
       #AUX_rgtSendBuffer.dLung := 0;
       #AUX_rgtSendBuffer.dID := #AUX_rgtSendBuffer.dID + 1;
       #AUX_rgtSendBuffer.dThick_um := #INO_tTrack.tLastPlacedCap.dThick_cmm;
   //    WRITE_BIG(src_variable := _byte_in_, dest_array := _variant_inout_, pos := _dint_inout_);
       #TMP_dPos := 0;
       #TMP_iRetVal:= WRITE_LITTLE(src_variable :=  #AUX_rgtSendBuffer.dLung, dest_array :=  #AUX_rgtSendBuffer_LittleEndian, pos := #TMP_dPos);
       #TMP_dPos := 4;
       #TMP_iRetVal := WRITE_LITTLE(src_variable := #AUX_rgtSendBuffer.dID, dest_array := #AUX_rgtSendBuffer_LittleEndian, pos := #TMP_dPos);
       #TMP_dPos := 8;
       #TMP_iRetVal := WRITE_LITTLE(src_variable := #AUX_rgtSendBuffer.dThick_um, dest_array := #AUX_rgtSendBuffer_LittleEndian, pos := #TMP_dPos);
       #AUX_dNumByteToSend := 0;
   END_IF;
END_REGION

REGION Network 25: ### SEND DATA TO CAMERA
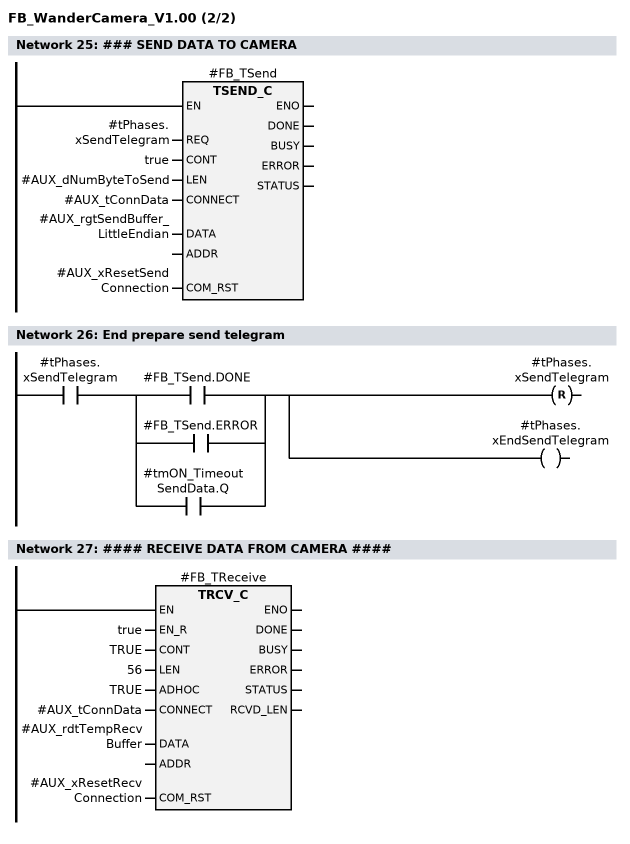
   #FB_TSend(REQ := #tPhases.xSendTelegram,   // TSEND_C
             CONT := true,
             LEN := #AUX_dNumByteToSend,
             CONNECT := #AUX_tConnData,
             DATA := #AUX_rgtSendBuffer_LittleEndian,
             COM_RST := #AUX_xResetSendConnection);
END_REGION

REGION Network 26: End prepare send telegram
   RUNG wire#powerrail
      Contact( #tPhases.xSendTelegram )
      wire#w1
      Contact( #FB_TSend.DONE )
      wire#w2
      R_Coil( #tPhases.xSendTelegram )
   END_RUNG
   RUNG wire#w1
      Contact( #FB_TSend.ERROR )
   END_RUNG wire#w2
   RUNG wire#w1
      Contact( #tmON_TimeoutSendData.Q )
   END_RUNG wire#w2
   RUNG wire#w2
      Coil( #tPhases.xEndSendTelegram )
   END_RUNG
   // the same network as SCL:
   #_w1 := #tPhases.xSendTelegram AND (#FB_TSend.DONE OR #FB_TSend.ERROR OR #tmON_TimeoutSendData.Q);
   IF #_w1 THEN #tPhases.xSendTelegram := FALSE; END_IF;
   #tPhases.xEndSendTelegram := #_w1;
END_REGION

REGION Network 27: #### RECEIVE DATA FROM CAMERA ####
   #FB_TReceive(EN_R := true,   // TRCV_C
                CONT := TRUE,
                LEN := 56,
                ADHOC := TRUE,
                CONNECT := #AUX_tConnData,
                DATA := #AUX_rdtTempRecvBuffer,
                COM_RST := #AUX_xResetRecvConnection);
END_REGION

REGION Network 28 (SCL): Manage data received
   IF #FB_TReceive.DONE THEN

       IF #FB_TReceive.RCVD_LEN > 0 THEN
           #TMP_dPos := 0;
           #TMP_iRetVal:= READ_LITTLE(src_array:=#AUX_rdtTempRecvBuffer, dest_Variable=>#AUX_rdtRecvBuffer.dLung, pos:=#TMP_dPos);
           #TMP_dPos := 4;
           #TMP_iRetVal := READ_LITTLE(src_array := #AUX_rdtTempRecvBuffer, dest_Variable => #AUX_rdtRecvBuffer.dID, pos := #TMP_dPos);
           #TMP_dPos := 8;
           #TMP_iRetVal := READ_LITTLE(src_array := #AUX_rdtTempRecvBuffer, dest_Variable => #AUX_rdtRecvBuffer.dTime1, pos := #TMP_dPos);
           #TMP_dPos := 12;
           #TMP_iRetVal := READ_LITTLE(src_array := #AUX_rdtTempRecvBuffer, dest_Variable => #AUX_rdtRecvBuffer.dTime2, pos := #TMP_dPos);
           #TMP_dPos := 16;
           #TMP_iRetVal := READ_LITTLE(src_array := #AUX_rdtTempRecvBuffer, dest_Variable => #AUX_rdtRecvBuffer.dStato, pos := #TMP_dPos);
           #TMP_dPos := 20;
           #TMP_iRetVal := READ_LITTLE(src_array := #AUX_rdtTempRecvBuffer, dest_Variable => #AUX_rdtRecvBuffer.dGrossZeroSide_um, pos := #TMP_dPos);
           #TMP_dPos := 24;
           #TMP_iRetVal := READ_LITTLE(src_array := #AUX_rdtTempRecvBuffer, dest_Variable => #AUX_rdtRecvBuffer.dNetExtZeroSide_um, pos := #TMP_dPos);
           #TMP_dPos := 28;
           #TMP_iRetVal := READ_LITTLE(src_array := #AUX_rdtTempRecvBuffer, dest_Variable => #AUX_rdtRecvBuffer.dNetCenterZeroSide_um, pos := #TMP_dPos);
           #TMP_dPos := 32;
           #TMP_iRetVal := READ_LITTLE(src_array := #AUX_rdtTempRecvBuffer, dest_Variable => #AUX_rdtRecvBuffer.dNetZeroSide_um, pos := #TMP_dPos);
           #TMP_dPos := 36;
           #TMP_iRetVal := READ_LITTLE(src_array := #AUX_rdtTempRecvBuffer, dest_Variable => #AUX_rdtRecvBuffer.dGrossOppSide_um, pos := #TMP_dPos);
           #TMP_dPos := 40;
           #TMP_iRetVal := READ_LITTLE(src_array := #AUX_rdtTempRecvBuffer, dest_Variable => #AUX_rdtRecvBuffer.dNetExtOppoSide_um, pos := #TMP_dPos);
           #TMP_dPos := 44;
           #TMP_iRetVal := READ_LITTLE(src_array := #AUX_rdtTempRecvBuffer, dest_Variable => #AUX_rdtRecvBuffer.dNetCenterOppoSide_um, pos := #TMP_dPos);
           #TMP_dPos := 48;
           #TMP_iRetVal := READ_LITTLE(src_array := #AUX_rdtTempRecvBuffer, dest_Variable => #AUX_rdtRecvBuffer.dNetOppoSide_um, pos := #TMP_dPos);
           #TMP_dPos := 52;
           #TMP_iRetVal := READ_LITTLE(src_array := #AUX_rdtTempRecvBuffer, dest_Variable => #AUX_rdtRecvBuffer.dLength, pos := #TMP_dPos);

           #OS_xNewDataAvailable := 1;
           #INO_tRibbon.rgtGlassData[#IN_dGlassDataMachineIndex].dDistSnapRoll_cmm := #tHMR.dDistanceFromSnaproll_cmm;

           //Update the position
           IF NOT #INO_tRibbon.rgtGlassDataUpdate[#IN_dGlassDataMachineIndex].xUpdateRequest THEN
               #INO_tRibbon.rgtGlassDataUpdate[#IN_dGlassDataMachineIndex].tData.dGrossWander_cmm := #tHMR.dCurrentGrossWander_cmm;
               #INO_tRibbon.rgtGlassDataUpdate[#IN_dGlassDataMachineIndex].tData.dNetWander_cmm := #tHMR.dCurrentNetWander_cmm;
               #INO_tRibbon.rgtGlassDataUpdate[#IN_dGlassDataMachineIndex].tData.dGrossWidth_cmm := #tHMR.dCurrentGrossWidth_cmm;
               #INO_tRibbon.rgtGlassDataUpdate[#IN_dGlassDataMachineIndex].tData.dNetWidth_cmm := #tHMR.dCurrentNetWidth_cmm;
               #INO_tRibbon.rgtGlassDataUpdate[#IN_dGlassDataMachineIndex].xUpdateRequest := TRUE;
           END_IF;
       END_IF;

   END_IF;
END_REGION

REGION Network 29 (SCL): Phase in progress
   GATHER(IN:=#tPhases,
          OUT=>#TMP_dwValue);

   IF #TMP_dwValue <> 0 THEN
       #ST_xPhaseProgr := TRUE;
   ELSE
       #ST_xPhaseProgr := FALSE;
   END_IF;
END_REGION
END_FUNCTION_BLOCK

// folder: 03_Programs_Logics/MCC1201/09_Zone

FUNCTION "ZUPS_Faults" : Void   // FC15, LAD
{ S7_Optimized_Access := 'TRUE' }
VERSION : 0.1
   VAR_TEMP
      TMP_dwValue : DWord;
   END_VAR
BEGIN

REGION Network 1 (SCL): Reset alarms
   IF "ZUPS".tmOFF_ResetAlarm.OUT_xDone THEN

       #TMP_dwValue := 0;

       SCATTER(IN := #TMP_dwValue,
               OUT => "DB_ZUPS_HMI".tAlm.tE);

       SCATTER(IN := #TMP_dwValue,
               OUT => "DB_ZUPS_HMI".tAlm.tS);

       SCATTER(IN := #TMP_dwValue,
               OUT => "DB_ZUPS_HMI".tAlm.tF);

       SCATTER(IN := #TMP_dwValue,
               OUT => "DB_ZUPS_HMI".tAlm.tW);

   END_IF;
END_REGION

REGION Network 2: Anomalies
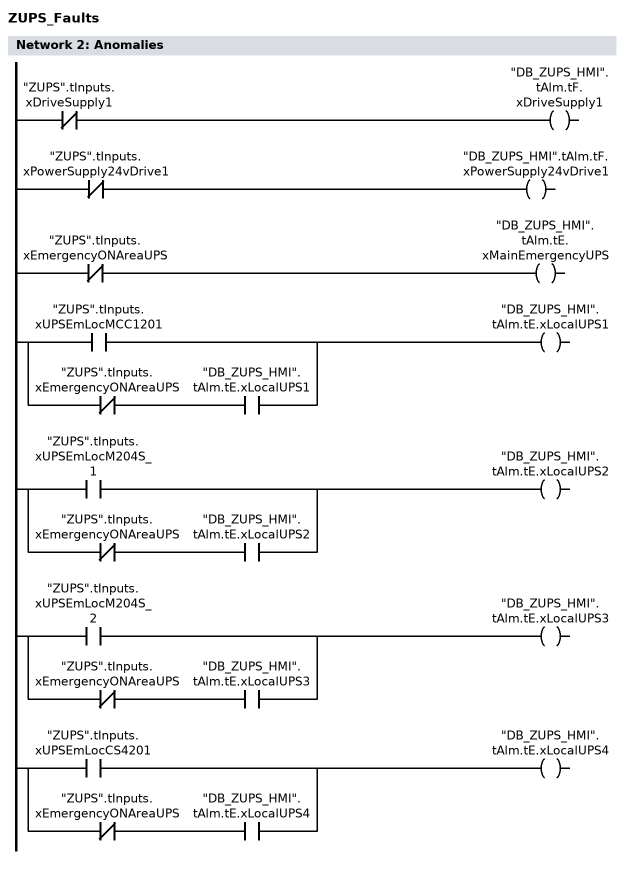
   RUNG wire#powerrail
      I_Contact( "ZUPS".tInputs.xDriveSupply1 )
      Coil( "DB_ZUPS_HMI".tAlm.tF.xDriveSupply1 )
   END_RUNG
   RUNG wire#powerrail
      I_Contact( "ZUPS".tInputs.xPowerSupply24vDrive1 )
      Coil( "DB_ZUPS_HMI".tAlm.tF.xPowerSupply24vDrive1 )
   END_RUNG
   RUNG wire#powerrail
      I_Contact( "ZUPS".tInputs.xEmergencyONAreaUPS )
      Coil( "DB_ZUPS_HMI".tAlm.tE.xMainEmergencyUPS )
   END_RUNG
   RUNG wire#powerrail
      Contact( "ZUPS".tInputs.xUPSEmLocMCC1201 )
      wire#w1
      Coil( "DB_ZUPS_HMI".tAlm.tE.xLocalUPS1 )
   END_RUNG
   RUNG wire#powerrail
      I_Contact( "ZUPS".tInputs.xEmergencyONAreaUPS )
      Contact( "DB_ZUPS_HMI".tAlm.tE.xLocalUPS1 )
   END_RUNG wire#w1
   RUNG wire#powerrail
      Contact( "ZUPS".tInputs.xUPSEmLocM204S_1 )
      wire#w2
      Coil( "DB_ZUPS_HMI".tAlm.tE.xLocalUPS2 )
   END_RUNG
   RUNG wire#powerrail
      I_Contact( "ZUPS".tInputs.xEmergencyONAreaUPS )
      Contact( "DB_ZUPS_HMI".tAlm.tE.xLocalUPS2 )
   END_RUNG wire#w2
   RUNG wire#powerrail
      Contact( "ZUPS".tInputs.xUPSEmLocM204S_2 )
      wire#w3
      Coil( "DB_ZUPS_HMI".tAlm.tE.xLocalUPS3 )
   END_RUNG
   RUNG wire#powerrail
      I_Contact( "ZUPS".tInputs.xEmergencyONAreaUPS )
      Contact( "DB_ZUPS_HMI".tAlm.tE.xLocalUPS3 )
   END_RUNG wire#w3
   RUNG wire#powerrail
      Contact( "ZUPS".tInputs.xUPSEmLocCS4201 )
      wire#w4
      Coil( "DB_ZUPS_HMI".tAlm.tE.xLocalUPS4 )
   END_RUNG
   RUNG wire#powerrail
      I_Contact( "ZUPS".tInputs.xEmergencyONAreaUPS )
      Contact( "DB_ZUPS_HMI".tAlm.tE.xLocalUPS4 )
   END_RUNG wire#w4
   // the same network as SCL:
   "DB_ZUPS_HMI".tAlm.tF.xDriveSupply1 := NOT "ZUPS".tInputs.xDriveSupply1;
   "DB_ZUPS_HMI".tAlm.tF.xPowerSupply24vDrive1 := NOT "ZUPS".tInputs.xPowerSupply24vDrive1;
   "DB_ZUPS_HMI".tAlm.tE.xMainEmergencyUPS := NOT "ZUPS".tInputs.xEmergencyONAreaUPS;
   "DB_ZUPS_HMI".tAlm.tE.xLocalUPS1 := "ZUPS".tInputs.xUPSEmLocMCC1201 OR (NOT "ZUPS".tInputs.xEmergencyONAreaUPS AND "DB_ZUPS_HMI".tAlm.tE.xLocalUPS1);
   "DB_ZUPS_HMI".tAlm.tE.xLocalUPS2 := "ZUPS".tInputs.xUPSEmLocM204S_1 OR (NOT "ZUPS".tInputs.xEmergencyONAreaUPS AND "DB_ZUPS_HMI".tAlm.tE.xLocalUPS2);
   "DB_ZUPS_HMI".tAlm.tE.xLocalUPS3 := "ZUPS".tInputs.xUPSEmLocM204S_2 OR (NOT "ZUPS".tInputs.xEmergencyONAreaUPS AND "DB_ZUPS_HMI".tAlm.tE.xLocalUPS3);
   "DB_ZUPS_HMI".tAlm.tE.xLocalUPS4 := "ZUPS".tInputs.xUPSEmLocCS4201 OR (NOT "ZUPS".tInputs.xEmergencyONAreaUPS AND "DB_ZUPS_HMI".tAlm.tE.xLocalUPS4);
END_REGION

REGION Network 3 (SCL): Calculate comulative status
   GATHER(IN:="DB_ZUPS_HMI".tAlm.tE,
              OUT=>#TMP_dwValue);

       IF "DB_ZUPS_HMI".tAlm.tE.xMainEmergencyUPS THEN
       "ZUPS".ST_xZoneEmergency := TRUE;
   ELSE
       "ZUPS".ST_xZoneEmergency := FALSE;
   END_IF;

   GATHER(IN:="DB_ZUPS_HMI".tAlm.tS,
              OUT=>#TMP_dwValue);

   IF #TMP_dwValue <> 0 THEN
       "ZUPS".ST_xZoneStoppingFaults := TRUE;
   ELSE
       "ZUPS".ST_xZoneStoppingFaults := FALSE;
   END_IF;

   GATHER(IN:="DB_ZUPS_HMI".tAlm.tF,
              OUT=>#TMP_dwValue);

   IF #TMP_dwValue <> 0 THEN
       "ZUPS".ST_xZoneFaults := TRUE;
   ELSE
       "ZUPS".ST_xZoneFaults := FALSE;
   END_IF;

   GATHER(IN:="DB_ZUPS_HMI".tAlm.tW,
              OUT=>#TMP_dwValue);

   IF #TMP_dwValue <> 0 THEN
       "ZUPS".ST_xZoneWarnings := TRUE;
   ELSE
       "ZUPS".ST_xZoneWarnings := FALSE;
   END_IF;

   IF "ZUPS".ST_xZoneEmergency AND "ZUPS".ST_xZoneStoppingFaults AND "ZUPS".ST_xZoneFaults THEN
       "ZUPS".ST_xZoneError := TRUE;
   ELSE
       "ZUPS".ST_xZoneError := FALSE;
   END_IF;
END_REGION
END_FUNCTION

FUNCTION "ZUPS_Logics" : Void   // FC17, LAD
{ S7_Optimized_Access := 'TRUE' }
VERSION : 0.1
   VAR_TEMP
      TMP_rlVal : LReal;
   END_VAR
   VAR_TEMP   // added for the SCL form of the ladder/FBD networks
      _w1 : Bool;
      _w2 : Bool;
   END_VAR
BEGIN

REGION Network 1: #### CONSTANTS ####
END_REGION

REGION Network 2 (SCL): ### SIMULATION ###
   IF "SIMULATION_ACTIVE" THEN
       "ZUPS".tInputs.xDriveSupply1 := TRUE;
       "ZUPS".tInputs.xPowerSupply24vDrive1 := TRUE; 
       "ZUPS".tInputs.xEmergencyONAreaUPS := true;

   END_IF;
END_REGION

REGION Network 3: #### MATCH ####
END_REGION

REGION Network 4: Emergency UPS OK delayed
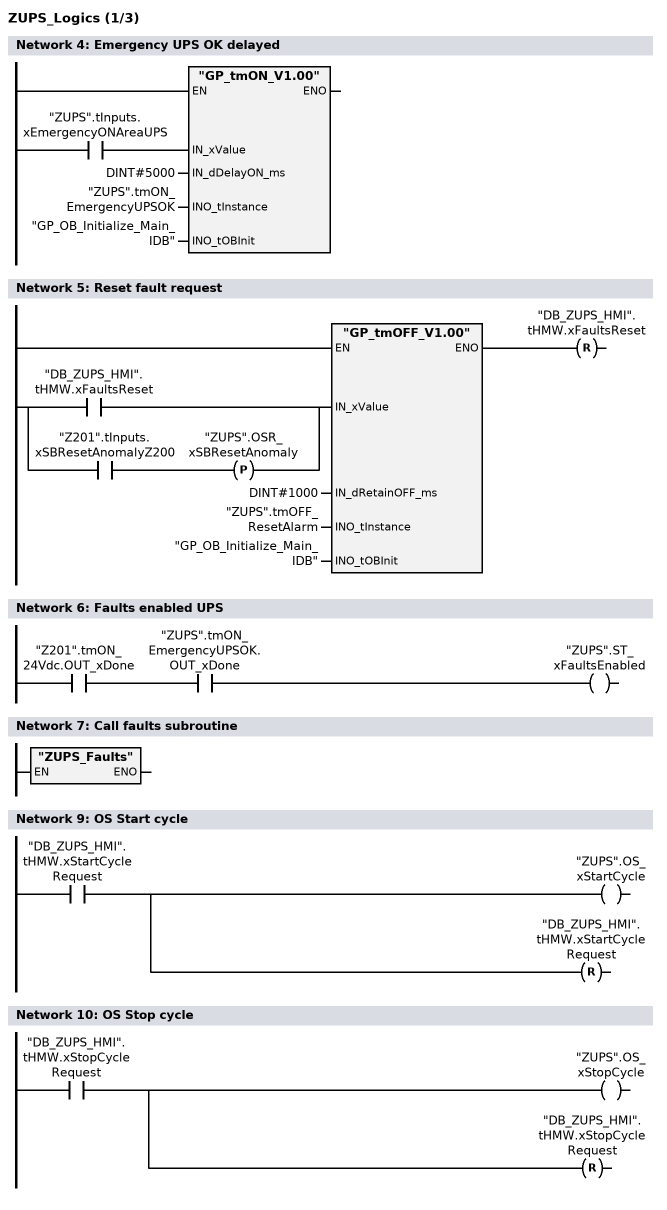
   RUNG wire#powerrail
      "GP_tmON_V1.00"(IN_xValue := wire#w1, IN_dDelayON_ms := DINT#5000, INO_tInstance := "ZUPS".tmON_EmergencyUPSOK, INO_tOBInit := "GP_OB_Initialize_Main_IDB")
   END_RUNG
   RUNG wire#powerrail
      Contact( "ZUPS".tInputs.xEmergencyONAreaUPS )
   END_RUNG wire#w1
   // the same network as SCL:
   "GP_tmON_V1.00"(IN_xValue := "ZUPS".tInputs.xEmergencyONAreaUPS,
                   IN_dDelayON_ms := DINT#5000,
                   INO_tInstance := "ZUPS".tmON_EmergencyUPSOK,
                   INO_tOBInit := "GP_OB_Initialize_Main_IDB");
END_REGION

REGION Network 5: Reset fault request
   RUNG wire#powerrail
      "GP_tmOFF_V1.00"(IN_xValue := wire#w1, IN_dRetainOFF_ms := DINT#1000, INO_tInstance := "ZUPS".tmOFF_ResetAlarm, INO_tOBInit := "GP_OB_Initialize_Main_IDB")
      R_Coil( "DB_ZUPS_HMI".tHMW.xFaultsReset )
   END_RUNG
   RUNG wire#powerrail
      Contact( "DB_ZUPS_HMI".tHMW.xFaultsReset )
   END_RUNG wire#w1
   RUNG wire#powerrail
      Contact( "Z201".tInputs.xSBResetAnomalyZ200 )
      P_Trig( "ZUPS".OSR_xSBResetAnomaly )
   END_RUNG wire#w1
   // the same network as SCL:
   #_w1 := "Z201".tInputs.xSBResetAnomalyZ200 AND NOT "ZUPS".OSR_xSBResetAnomaly;   // rising edge
   "ZUPS".OSR_xSBResetAnomaly := "Z201".tInputs.xSBResetAnomalyZ200;
   "GP_tmOFF_V1.00"(IN_xValue := "DB_ZUPS_HMI".tHMW.xFaultsReset OR #_w1,
                    IN_dRetainOFF_ms := DINT#1000,
                    INO_tInstance := "ZUPS".tmOFF_ResetAlarm,
                    INO_tOBInit := "GP_OB_Initialize_Main_IDB",
                    ENO => #_w2);
   IF #_w2 THEN "DB_ZUPS_HMI".tHMW.xFaultsReset := FALSE; END_IF;
END_REGION

REGION Network 6: Faults enabled UPS
   RUNG wire#powerrail
      Contact( "Z201".tmON_24Vdc.OUT_xDone )
      Contact( "ZUPS".tmON_EmergencyUPSOK.OUT_xDone )
      Coil( "ZUPS".ST_xFaultsEnabled )
   END_RUNG
   // the same network as SCL:
   "ZUPS".ST_xFaultsEnabled := "Z201".tmON_24Vdc.OUT_xDone AND "ZUPS".tmON_EmergencyUPSOK.OUT_xDone;
END_REGION

REGION Network 7: Call faults subroutine
   RUNG wire#powerrail
      "ZUPS_Faults"()
   END_RUNG
   // the same network as SCL:
   "ZUPS_Faults"();
END_REGION

REGION Network 8: #### START/STOP ZONE ####
END_REGION

REGION Network 9: OS Start cycle
   RUNG wire#powerrail
      Contact( "DB_ZUPS_HMI".tHMW.xStartCycleRequest )
      wire#w1
      Coil( "ZUPS".OS_xStartCycle )
   END_RUNG
   RUNG wire#w1
      R_Coil( "DB_ZUPS_HMI".tHMW.xStartCycleRequest )
   END_RUNG
   // the same network as SCL:
   "ZUPS".OS_xStartCycle := "DB_ZUPS_HMI".tHMW.xStartCycleRequest;
   IF "DB_ZUPS_HMI".tHMW.xStartCycleRequest THEN "DB_ZUPS_HMI".tHMW.xStartCycleRequest := FALSE; END_IF;
END_REGION

REGION Network 10: OS Stop cycle
   RUNG wire#powerrail
      Contact( "DB_ZUPS_HMI".tHMW.xStopCycleRequest )
      wire#w1
      Coil( "ZUPS".OS_xStopCycle )
   END_RUNG
   RUNG wire#w1
      R_Coil( "DB_ZUPS_HMI".tHMW.xStopCycleRequest )
   END_RUNG
   // the same network as SCL:
   "ZUPS".OS_xStopCycle := "DB_ZUPS_HMI".tHMW.xStopCycleRequest;
   IF "DB_ZUPS_HMI".tHMW.xStopCycleRequest THEN "DB_ZUPS_HMI".tHMW.xStopCycleRequest := FALSE; END_IF;
END_REGION

REGION Network 11: OS Force stop cycle
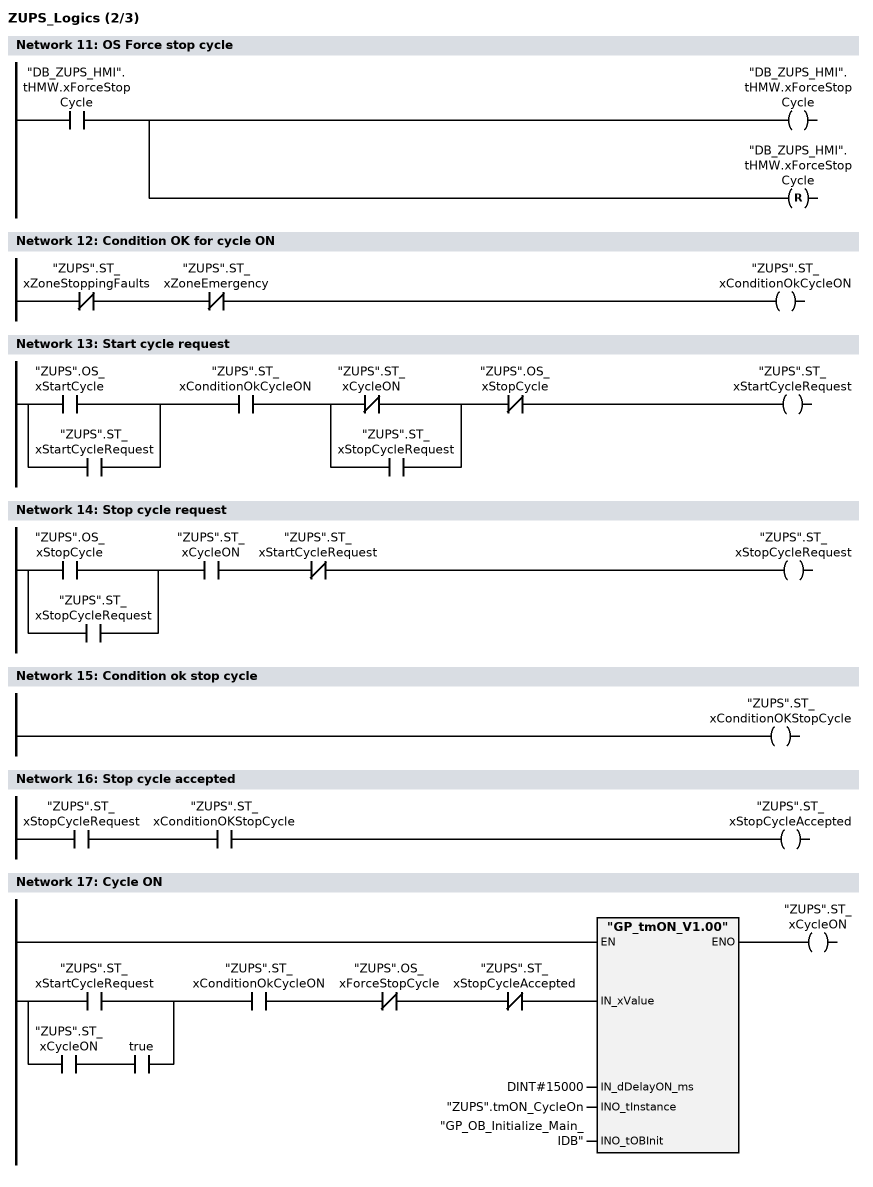
   RUNG wire#powerrail
      Contact( "DB_ZUPS_HMI".tHMW.xForceStopCycle )
      wire#w1
      Coil( "DB_ZUPS_HMI".tHMW.xForceStopCycle )
   END_RUNG
   RUNG wire#w1
      R_Coil( "DB_ZUPS_HMI".tHMW.xForceStopCycle )
   END_RUNG
   // the same network as SCL:
   #_w1 := "DB_ZUPS_HMI".tHMW.xForceStopCycle;
   "DB_ZUPS_HMI".tHMW.xForceStopCycle := "DB_ZUPS_HMI".tHMW.xForceStopCycle;
   IF #_w1 THEN "DB_ZUPS_HMI".tHMW.xForceStopCycle := FALSE; END_IF;
END_REGION

REGION Network 12: Condition OK for cycle ON
   RUNG wire#powerrail
      I_Contact( "ZUPS".ST_xZoneStoppingFaults )
      I_Contact( "ZUPS".ST_xZoneEmergency )
      Coil( "ZUPS".ST_xConditionOkCycleON )
   END_RUNG
   // the same network as SCL:
   "ZUPS".ST_xConditionOkCycleON := NOT "ZUPS".ST_xZoneStoppingFaults AND NOT "ZUPS".ST_xZoneEmergency;
END_REGION

REGION Network 13: Start cycle request
   RUNG wire#powerrail
      Contact( "ZUPS".OS_xStartCycle )
      wire#w1
      Contact( "ZUPS".ST_xConditionOkCycleON )
      wire#w2
      I_Contact( "ZUPS".ST_xCycleON )
      wire#w3
      I_Contact( "ZUPS".OS_xStopCycle )
      Coil( "ZUPS".ST_xStartCycleRequest )
   END_RUNG
   RUNG wire#powerrail
      Contact( "ZUPS".ST_xStartCycleRequest )
   END_RUNG wire#w1
   RUNG wire#w2
      Contact( "ZUPS".ST_xStopCycleRequest )
   END_RUNG wire#w3
   // the same network as SCL:
   "ZUPS".ST_xStartCycleRequest := ("ZUPS".OS_xStartCycle OR "ZUPS".ST_xStartCycleRequest) AND "ZUPS".ST_xConditionOkCycleON AND (NOT "ZUPS".ST_xCycleON OR "ZUPS".ST_xStopCycleRequest) AND NOT "ZUPS".OS_xStopCycle;
END_REGION

REGION Network 14: Stop cycle request
   RUNG wire#powerrail
      Contact( "ZUPS".OS_xStopCycle )
      wire#w1
      Contact( "ZUPS".ST_xCycleON )
      I_Contact( "ZUPS".ST_xStartCycleRequest )
      Coil( "ZUPS".ST_xStopCycleRequest )
   END_RUNG
   RUNG wire#powerrail
      Contact( "ZUPS".ST_xStopCycleRequest )
   END_RUNG wire#w1
   // the same network as SCL:
   "ZUPS".ST_xStopCycleRequest := ("ZUPS".OS_xStopCycle OR "ZUPS".ST_xStopCycleRequest) AND "ZUPS".ST_xCycleON AND NOT "ZUPS".ST_xStartCycleRequest;
END_REGION

REGION Network 15: Condition ok stop cycle
   RUNG wire#powerrail
      Coil( "ZUPS".ST_xConditionOKStopCycle )
   END_RUNG
   // the same network as SCL:
   "ZUPS".ST_xConditionOKStopCycle := TRUE;
END_REGION

REGION Network 16: Stop cycle accepted
   RUNG wire#powerrail
      Contact( "ZUPS".ST_xStopCycleRequest )
      Contact( "ZUPS".ST_xConditionOKStopCycle )
      Coil( "ZUPS".ST_xStopCycleAccepted )
   END_RUNG
   // the same network as SCL:
   "ZUPS".ST_xStopCycleAccepted := "ZUPS".ST_xStopCycleRequest AND "ZUPS".ST_xConditionOKStopCycle;
END_REGION

REGION Network 17: Cycle ON
   RUNG wire#powerrail
      "GP_tmON_V1.00"(IN_xValue := wire#w2, IN_dDelayON_ms := DINT#15000, INO_tInstance := "ZUPS".tmON_CycleOn, INO_tOBInit := "GP_OB_Initialize_Main_IDB")
      Coil( "ZUPS".ST_xCycleON )
   END_RUNG
   RUNG wire#powerrail
      Contact( "ZUPS".ST_xStartCycleRequest )
      wire#w1
      Contact( "ZUPS".ST_xConditionOkCycleON )
      I_Contact( "ZUPS".OS_xForceStopCycle )
      I_Contact( "ZUPS".ST_xStopCycleAccepted )
   END_RUNG wire#w2
   RUNG wire#powerrail
      Contact( "ZUPS".ST_xCycleON )
      Contact( true )
   END_RUNG wire#w1
   // the same network as SCL:
   "GP_tmON_V1.00"(IN_xValue := ("ZUPS".ST_xStartCycleRequest OR ("ZUPS".ST_xCycleON AND true)) AND "ZUPS".ST_xConditionOkCycleON AND NOT "ZUPS".OS_xForceStopCycle AND NOT "ZUPS".ST_xStopCycleAccepted,
                   IN_dDelayON_ms := DINT#15000,
                   INO_tInstance := "ZUPS".tmON_CycleOn,
                   INO_tOBInit := "GP_OB_Initialize_Main_IDB",
                   ENO => #_w1);
   "ZUPS".ST_xCycleON := #_w1;
END_REGION

REGION Network 18: Cycle ON delayed
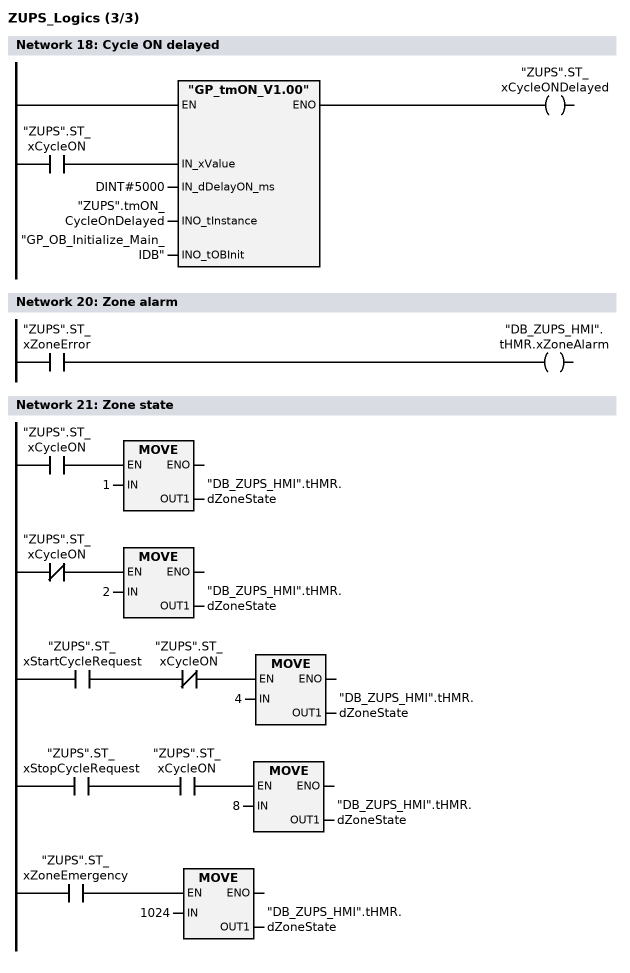
   RUNG wire#powerrail
      "GP_tmON_V1.00"(IN_xValue := wire#w1, IN_dDelayON_ms := DINT#5000, INO_tInstance := "ZUPS".tmON_CycleOnDelayed, INO_tOBInit := "GP_OB_Initialize_Main_IDB")
      Coil( "ZUPS".ST_xCycleONDelayed )
   END_RUNG
   RUNG wire#powerrail
      Contact( "ZUPS".ST_xCycleON )
   END_RUNG wire#w1
   // the same network as SCL:
   "GP_tmON_V1.00"(IN_xValue := "ZUPS".ST_xCycleON,
                   IN_dDelayON_ms := DINT#5000,
                   INO_tInstance := "ZUPS".tmON_CycleOnDelayed,
                   INO_tOBInit := "GP_OB_Initialize_Main_IDB",
                   ENO => #_w1);
   "ZUPS".ST_xCycleONDelayed := #_w1;
END_REGION

REGION Network 19: #### HMI STATUSES ####
END_REGION

REGION Network 20: Zone alarm
   RUNG wire#powerrail
      Contact( "ZUPS".ST_xZoneError )
      Coil( "DB_ZUPS_HMI".tHMR.xZoneAlarm )
   END_RUNG
   // the same network as SCL:
   "DB_ZUPS_HMI".tHMR.xZoneAlarm := "ZUPS".ST_xZoneError;
END_REGION

REGION Network 21: Zone state
   RUNG wire#powerrail
      Contact( "ZUPS".ST_xCycleON )
      Move(in := 1, out1 => "DB_ZUPS_HMI".tHMR.dZoneState)
   END_RUNG
   RUNG wire#powerrail
      I_Contact( "ZUPS".ST_xCycleON )
      Move(in := 2, out1 => "DB_ZUPS_HMI".tHMR.dZoneState)
   END_RUNG
   RUNG wire#powerrail
      Contact( "ZUPS".ST_xStartCycleRequest )
      I_Contact( "ZUPS".ST_xCycleON )
      Move(in := 4, out1 => "DB_ZUPS_HMI".tHMR.dZoneState)
   END_RUNG
   RUNG wire#powerrail
      Contact( "ZUPS".ST_xStopCycleRequest )
      Contact( "ZUPS".ST_xCycleON )
      Move(in := 8, out1 => "DB_ZUPS_HMI".tHMR.dZoneState)
   END_RUNG
   RUNG wire#powerrail
      Contact( "ZUPS".ST_xZoneEmergency )
      Move(in := 1024, out1 => "DB_ZUPS_HMI".tHMR.dZoneState)
   END_RUNG
   // the same network as SCL:
   IF "ZUPS".ST_xCycleON THEN "DB_ZUPS_HMI".tHMR.dZoneState := 1; END_IF;
   IF NOT "ZUPS".ST_xCycleON THEN "DB_ZUPS_HMI".tHMR.dZoneState := 2; END_IF;
   IF "ZUPS".ST_xStartCycleRequest AND NOT "ZUPS".ST_xCycleON THEN
       "DB_ZUPS_HMI".tHMR.dZoneState := 4;
   END_IF;
   IF "ZUPS".ST_xStopCycleRequest AND "ZUPS".ST_xCycleON THEN "DB_ZUPS_HMI".tHMR.dZoneState := 8; END_IF;
   IF "ZUPS".ST_xZoneEmergency THEN "DB_ZUPS_HMI".tHMR.dZoneState := 1024; END_IF;
END_REGION
END_FUNCTION

FUNCTION "ZUPS_Output" : Void   // FC28, LAD
{ S7_Optimized_Access := 'TRUE' }
VERSION : 0.1
BEGIN

REGION Network 1: HL emergency
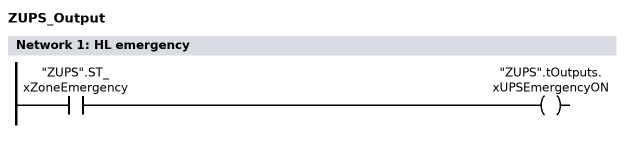
   RUNG wire#powerrail
      Contact( "ZUPS".ST_xZoneEmergency )
      Coil( "ZUPS".tOutputs.xUPSEmergencyON )
   END_RUNG
   // the same network as SCL:
   "ZUPS".tOutputs.xUPSEmergencyON := "ZUPS".ST_xZoneEmergency;
END_REGION
END_FUNCTION

FUNCTION "Z201_Logics" : Void   // FC29, LAD
{ S7_Optimized_Access := 'TRUE' }
VERSION : 0.1
   VAR_TEMP
      TMP_rlVal : LReal;
   END_VAR
   VAR_TEMP   // added for the SCL form of the ladder/FBD networks
      _w1 : Bool;
      _w2 : Bool;
   END_VAR
BEGIN

REGION Network 1: #### CONSTANTS ####
END_REGION

REGION Network 2 (SCL): ### SIMULATION ###
   IF "SIMULATION_ACTIVE" THEN

       "Z201".tInputs.xCPUAEnabled := TRUE;
       "Z201".tInputs.xCPUBEnabled := FALSE;
       "Z201".tInputs.xCPUARecognition := TRUE;
       "Z201".tInputs.xCPUBRecognition := FALSE;
       "Z201".tInputs.xM216FanFeedback := TRUE;

       "Z201".tInputs.xPowerSupply24vLogic1 := TRUE;
       "Z201".tInputs.xPowerSupply24vLogic2 := TRUE;
       "Z201".tInputs.xPowerSupply24vLogic3 := TRUE;
       "Z201".tInputs.xPowerSupply24vLogic4 := TRUE;
       "Z201".tInputs.xPowerSupply230vAux := TRUE;
       "Z201".tInputs.xPowerSuppluyOut24vUnderUpsEmOk := TRUE;
       "Z201".tInputs.xPowerSuppluyOut24vUnderEmOk := TRUE;
       "Z201".tInputs.xDriveSupply2 := TRUE;
       "Z201".tInputs.xPowerSupply24vDrive2 := TRUE;

       "Z201".tInputs.xMainEmergencyON := TRUE;
   END_IF;
   "TestTag64" := 0;
   "TestTag64".%X40 := 1;
END_REGION

REGION Network 3: #### MATCH ####
END_REGION

REGION Network 4: #### PLC ACTIVE ####
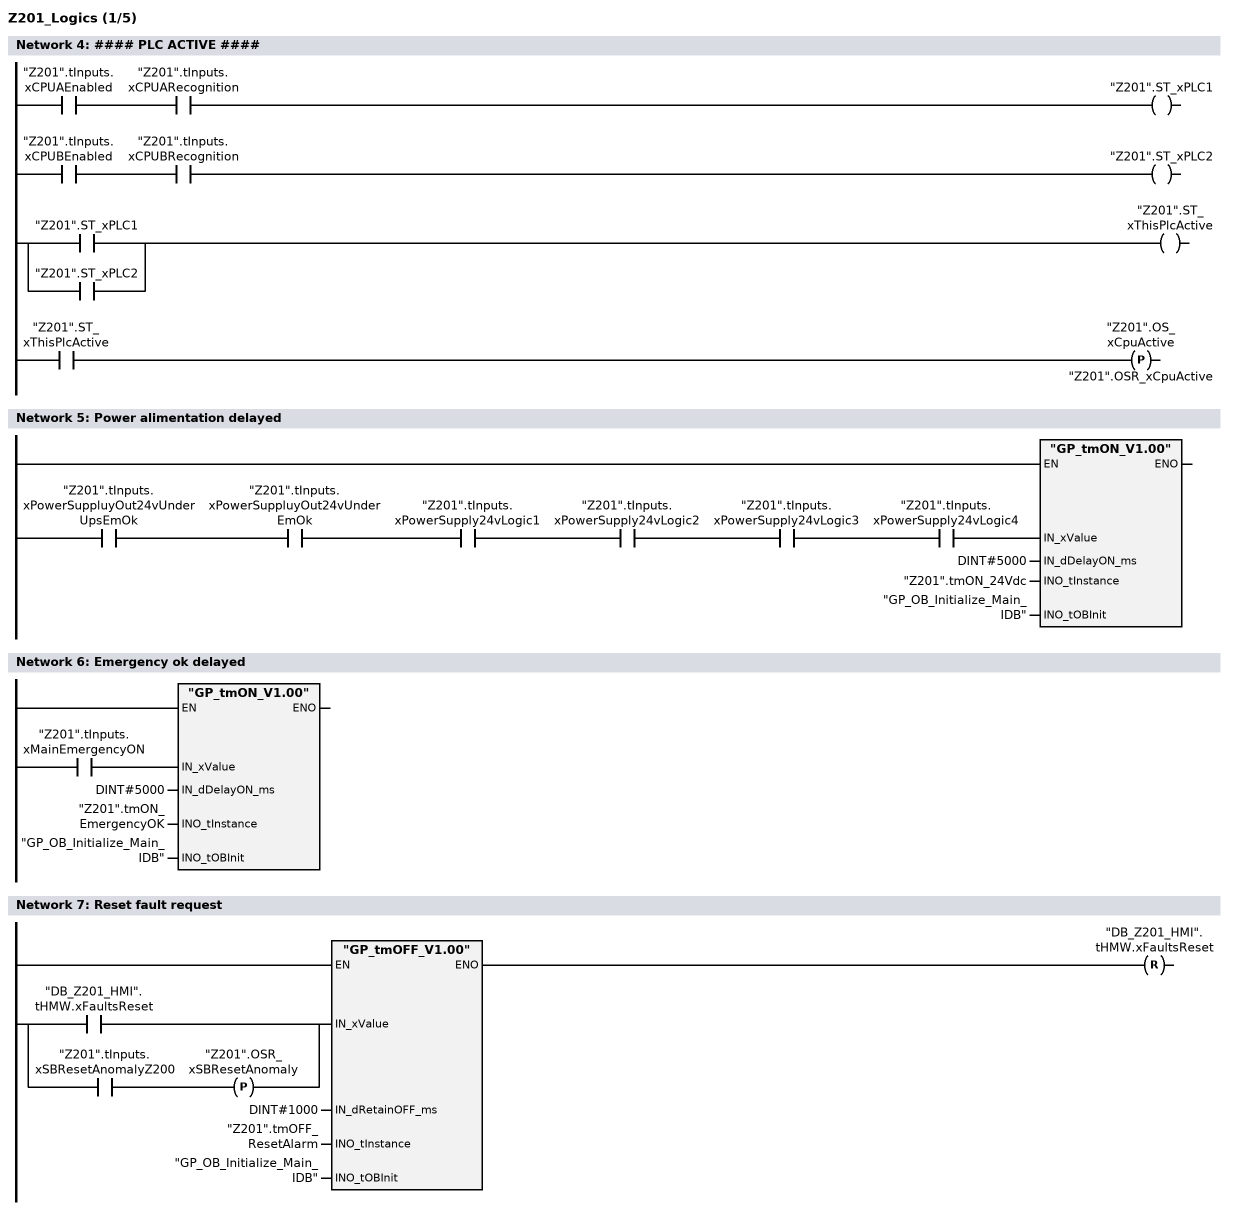
   "Z201".ST_xPLC1 := "Z201".tInputs.xCPUAEnabled AND "Z201".tInputs.xCPUARecognition;
   "Z201".ST_xPLC2 := "Z201".tInputs.xCPUBEnabled AND "Z201".tInputs.xCPUBRecognition;
   "Z201".ST_xThisPlcActive := "Z201".ST_xPLC1 OR "Z201".ST_xPLC2;
   "Z201".OS_xCpuActive := "Z201".ST_xThisPlcActive AND NOT "Z201".OSR_xCpuActive;   // rising edge
   "Z201".OSR_xCpuActive := "Z201".ST_xThisPlcActive;
END_REGION

REGION Network 5: Power alimentation delayed
   RUNG wire#powerrail
      "GP_tmON_V1.00"(IN_xValue := wire#w1, IN_dDelayON_ms := DINT#5000, INO_tInstance := "Z201".tmON_24Vdc, INO_tOBInit := "GP_OB_Initialize_Main_IDB")
   END_RUNG
   RUNG wire#powerrail
      Contact( "Z201".tInputs.xPowerSuppluyOut24vUnderUpsEmOk )
      Contact( "Z201".tInputs.xPowerSuppluyOut24vUnderEmOk )
      Contact( "Z201".tInputs.xPowerSupply24vLogic1 )
      Contact( "Z201".tInputs.xPowerSupply24vLogic2 )
      Contact( "Z201".tInputs.xPowerSupply24vLogic3 )
      Contact( "Z201".tInputs.xPowerSupply24vLogic4 )
   END_RUNG wire#w1
   // the same network as SCL:
   "GP_tmON_V1.00"(IN_xValue := "Z201".tInputs.xPowerSuppluyOut24vUnderUpsEmOk AND "Z201".tInputs.xPowerSuppluyOut24vUnderEmOk AND "Z201".tInputs.xPowerSupply24vLogic1 AND "Z201".tInputs.xPowerSupply24vLogic2 AND "Z201".tInputs.xPowerSupply24vLogic3 AND "Z201".tInputs.xPowerSupply24vLogic4,
                   IN_dDelayON_ms := DINT#5000,
                   INO_tInstance := "Z201".tmON_24Vdc,
                   INO_tOBInit := "GP_OB_Initialize_Main_IDB");
END_REGION

REGION Network 6: Emergency ok delayed
   RUNG wire#powerrail
      "GP_tmON_V1.00"(IN_xValue := wire#w1, IN_dDelayON_ms := DINT#5000, INO_tInstance := "Z201".tmON_EmergencyOK, INO_tOBInit := "GP_OB_Initialize_Main_IDB")
   END_RUNG
   RUNG wire#powerrail
      Contact( "Z201".tInputs.xMainEmergencyON )
   END_RUNG wire#w1
   // the same network as SCL:
   "GP_tmON_V1.00"(IN_xValue := "Z201".tInputs.xMainEmergencyON,
                   IN_dDelayON_ms := DINT#5000,
                   INO_tInstance := "Z201".tmON_EmergencyOK,
                   INO_tOBInit := "GP_OB_Initialize_Main_IDB");
END_REGION

REGION Network 7: Reset fault request
   RUNG wire#powerrail
      "GP_tmOFF_V1.00"(IN_xValue := wire#w1, IN_dRetainOFF_ms := DINT#1000, INO_tInstance := "Z201".tmOFF_ResetAlarm, INO_tOBInit := "GP_OB_Initialize_Main_IDB")
      R_Coil( "DB_Z201_HMI".tHMW.xFaultsReset )
   END_RUNG
   RUNG wire#powerrail
      Contact( "DB_Z201_HMI".tHMW.xFaultsReset )
   END_RUNG wire#w1
   RUNG wire#powerrail
      Contact( "Z201".tInputs.xSBResetAnomalyZ200 )
      P_Trig( "Z201".OSR_xSBResetAnomaly )
   END_RUNG wire#w1
   // the same network as SCL:
   #_w1 := "Z201".tInputs.xSBResetAnomalyZ200 AND NOT "Z201".OSR_xSBResetAnomaly;   // rising edge
   "Z201".OSR_xSBResetAnomaly := "Z201".tInputs.xSBResetAnomalyZ200;
   "GP_tmOFF_V1.00"(IN_xValue := "DB_Z201_HMI".tHMW.xFaultsReset OR #_w1,
                    IN_dRetainOFF_ms := DINT#1000,
                    INO_tInstance := "Z201".tmOFF_ResetAlarm,
                    INO_tOBInit := "GP_OB_Initialize_Main_IDB",
                    ENO => #_w2);
   IF #_w2 THEN "DB_Z201_HMI".tHMW.xFaultsReset := FALSE; END_IF;
END_REGION

REGION Network 8: General reset
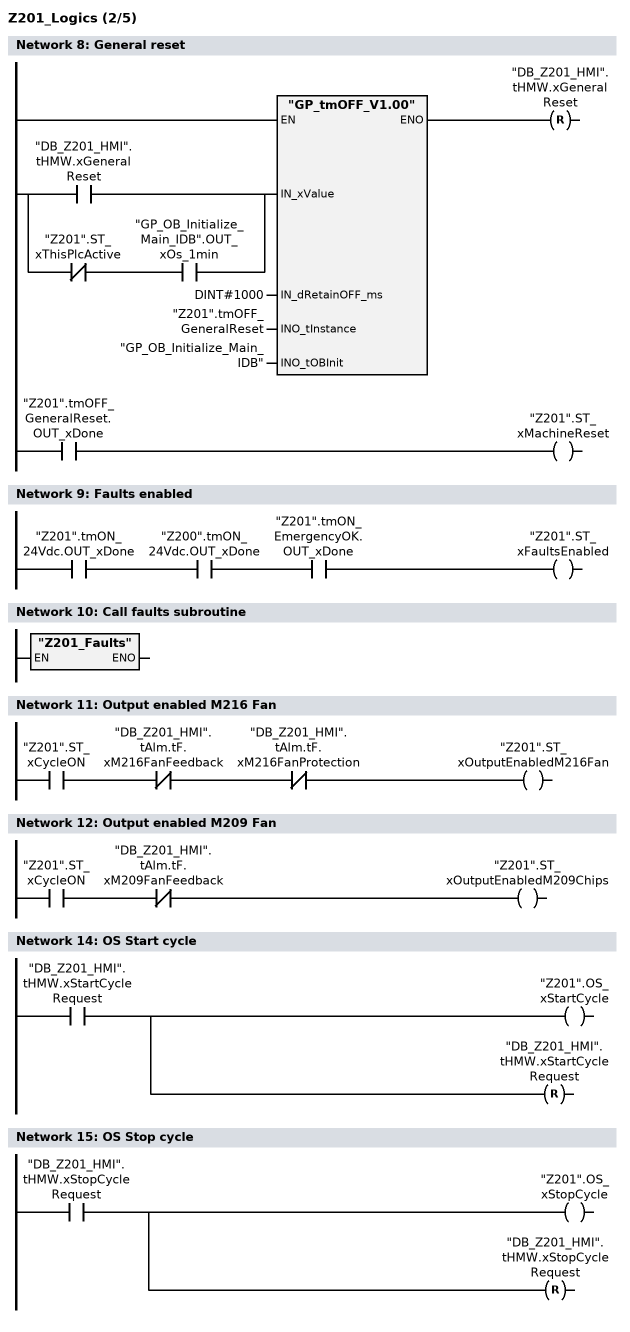
   RUNG wire#powerrail
      "GP_tmOFF_V1.00"(IN_xValue := wire#w1, IN_dRetainOFF_ms := DINT#1000, INO_tInstance := "Z201".tmOFF_GeneralReset, INO_tOBInit := "GP_OB_Initialize_Main_IDB")
      R_Coil( "DB_Z201_HMI".tHMW.xGeneralReset )
   END_RUNG
   RUNG wire#powerrail
      Contact( "DB_Z201_HMI".tHMW.xGeneralReset )
   END_RUNG wire#w1
   RUNG wire#powerrail
      I_Contact( "Z201".ST_xThisPlcActive )
      Contact( "GP_OB_Initialize_Main_IDB".OUT_xOs_1min )
   END_RUNG wire#w1
   RUNG wire#powerrail
      Contact( "Z201".tmOFF_GeneralReset.OUT_xDone )
      Coil( "Z201".ST_xMachineReset )
   END_RUNG
   // the same network as SCL:
   "GP_tmOFF_V1.00"(IN_xValue := "DB_Z201_HMI".tHMW.xGeneralReset OR (NOT "Z201".ST_xThisPlcActive AND "GP_OB_Initialize_Main_IDB".OUT_xOs_1min),
                    IN_dRetainOFF_ms := DINT#1000,
                    INO_tInstance := "Z201".tmOFF_GeneralReset,
                    INO_tOBInit := "GP_OB_Initialize_Main_IDB",
                    ENO => #_w1);
   IF #_w1 THEN "DB_Z201_HMI".tHMW.xGeneralReset := FALSE; END_IF;
   "Z201".ST_xMachineReset := "Z201".tmOFF_GeneralReset.OUT_xDone;
END_REGION

REGION Network 9: Faults enabled
   RUNG wire#powerrail
      Contact( "Z201".tmON_24Vdc.OUT_xDone )
      Contact( "Z200".tmON_24Vdc.OUT_xDone )
      Contact( "Z201".tmON_EmergencyOK.OUT_xDone )
      Coil( "Z201".ST_xFaultsEnabled )
   END_RUNG
   // the same network as SCL:
   "Z201".ST_xFaultsEnabled := "Z201".tmON_24Vdc.OUT_xDone AND "Z200".tmON_24Vdc.OUT_xDone AND "Z201".tmON_EmergencyOK.OUT_xDone;
END_REGION

REGION Network 10: Call faults subroutine
   RUNG wire#powerrail
      "Z201_Faults"()
   END_RUNG
   // the same network as SCL:
   "Z201_Faults"();
END_REGION

REGION Network 11: Output enabled M216 Fan
   RUNG wire#powerrail
      Contact( "Z201".ST_xCycleON )
      I_Contact( "DB_Z201_HMI".tAlm.tF.xM216FanFeedback )
      I_Contact( "DB_Z201_HMI".tAlm.tF.xM216FanProtection )
      Coil( "Z201".ST_xOutputEnabledM216Fan )
   END_RUNG
   // the same network as SCL:
   "Z201".ST_xOutputEnabledM216Fan := "Z201".ST_xCycleON AND NOT "DB_Z201_HMI".tAlm.tF.xM216FanFeedback AND NOT "DB_Z201_HMI".tAlm.tF.xM216FanProtection;
END_REGION
